   t[3580] := 1_070_001_024;
   t[3581] := 1_070_002_013;
   t[3582] := 1_070_003_096;
   t[3583] := 2_071_201_008;
   t[3584] := 2_071_202_005;
   t[3585] := 2_071_403_104;
   t[3586] := 71403105;
   t[3587] := 71502007;
   t[3588] := 71503043;
   t[3589] := 1_071_501_000;
   t[3590] := 1_071_502_003;
   t[3591] := 73603047;
   t[3592] := 2_073_602_002;
   t[3593] := 73602000;
   t[3594] := 73603013;
   t[3595] := 83001002;
   t[3596] := 1_083_001_014;
   t[3597] := 1_083_002_004;
   t[3598] := 1_084_801_030;
   t[3599] := 1_084_802_012;
   t[3600] := 2_084_801_022;
   t[3601] := 2_084_802_008;
   t[3602] := 84801020;
   t[3603] := 1_084_801_016;
   t[3604] := 85001000;
   t[3605] := 85002000;
   t[3606] := 2_085_101_016;
   t[3607] := 2_085_102_008;
   t[3608] := 1_086_312_107;
   t[3609] := 2_089_703_009;
   t[3610] := 2_090_203_001;
   t[3611] := 90203000;
   t[3612] := 94102009;
   t[3613] := 1_094_101_024;
   t[3614] := 1_094_102_013;
   t[3615] := 1_094_103_096;
   t[3616] := 1_095_201_008;
   t[3617] := 1_095_202_005;
   t[3618] := 2_095_403_104;
   t[3619] := 95403105;
   t[3620] := 95502007;
   t[3621] := 95503043;
   t[3622] := 1_095_501_000;
   t[3623] := 1_095_502_003;
   t[3624] := 97603047;
   t[3625] := 2_097_602_002;
   t[3626] := 97602000;
   t[3627] := 97603013;
   t[3628] := 1_110_312_108;
   t[3629] := 2_113_803_009;
   t[3630] := 114_303_001;
   t[3631] := 1_114_303_000;
   t[3632] := 148_701_002;
   t[3633] := 1_148_701_014;
   t[3634] := 1_148_702_004;
   t[3635] := 150_501_030;
   t[3636] := 150_502_012;
   t[3637] := 1_150_501_022;
   t[3638] := 1_150_502_008;
   t[3639] := 2_150_501_020;
   t[3640] := 150_501_016;
   t[3641] := 150_701_000;
   t[3642] := 150_702_000;
   t[3643] := 150_801_016;
   t[3644] := 150_802_008;
   t[3645] := 1_151_101_000;
   t[3646] := 1_151_102_000;
   t[3647] := 1_151_101_016;
   t[3648] := 1_151_102_008;
   t[3649] := 2_153_502_009;
   t[3650] := 153_501_024;
   t[3651] := 153_502_013;
   t[3652] := 153_503_096;
   t[3653] := 1_154_001_008;
   t[3654] := 1_154_002_005;
   t[3655] := 2_154_101_024;
   t[3656] := 2_154_102_013;
   t[3657] := 2_154_301_008;
   t[3658] := 2_154_302_005;
   t[3659] := 2_154_401_024;
   t[3660] := 2_154_402_013;
   t[3661] := 2_154_601_008;
   t[3662] := 2_154_602_005;
   t[3663] := 154_903_104;
   t[3664] := 1_154_903_105;
   t[3665] := 155_002_007;
   t[3666] := 155_003_043;
   t[3667] := 1_155_001_000;
   t[3668] := 1_155_002_003;
   t[3669] := 2_157_003_047;
   t[3670] := 1_157_002_002;
   t[3671] := 2_157_002_000;
   t[3672] := 2_157_003_013;
   t[3673] := 170_012_109;
   t[3674] := 2_173_703_009;
   t[3675] := 2_174_103_001;
   t[3676] := 174_103_000;
   t[3677] := 269_401_002;
   t[3678] := 1_269_401_014;
   t[3679] := 1_269_402_004;
   t[3680] := 271_101_030;
   t[3681] := 271_102_012;
   t[3682] := 1_271_101_022;
   t[3683] := 1_271_102_008;
   t[3684] := 2_271_101_020;
   t[3685] := 271_101_016;
   t[3686] := 1_271_301_000;
   t[3687] := 1_271_302_000;
   t[3688] := 2_271_401_016;
   t[3689] := 2_271_402_008;
   t[3690] := 274_102_009;
   t[3691] := 1_274_101_024;
   t[3692] := 1_274_102_013;
   t[3693] := 1_274_103_096;
   t[3694] := 2_275_101_008;
   t[3695] := 2_275_102_005;
   t[3696] := 1_275_403_104;
   t[3697] := 2_275_403_105;
   t[3698] := 1_275_402_007;
   t[3699] := 1_275_403_043;
   t[3700] := 2_275_401_000;
   t[3701] := 2_275_402_003;
   t[3702] := 2_277_403_047;
   t[3703] := 1_277_402_002;
   t[3704] := 2_277_402_000;
   t[3705] := 2_277_403_013;
   t[3706] := 1_290_212_110;
   t[3707] := 2_294_103_009;
   t[3708] := 294_303_001;
   t[3709] := 1_294_303_000;
   t[3710] := 380_401_002;
   t[3711] := 1_380_401_014;
   t[3712] := 1_380_402_004;
   t[3713] := 2_382_301_030;
   t[3714] := 2_382_302_012;
   t[3715] := 382_301_022;
   t[3716] := 382_302_008;
   t[3717] := 1_382_301_020;
   t[3718] := 2_382_301_016;
   t[3719] := 382_501_000;
   t[3720] := 382_502_000;
   t[3721] := 2_382_601_016;
   t[3722] := 2_382_602_008;
   t[3723] := 1_385_202_009;
   t[3724] := 2_385_201_024;
   t[3725] := 2_385_202_013;
   t[3726] := 2_385_203_096;
   t[3727] := 2_386_301_008;
   t[3728] := 2_386_302_005;
   t[3729] := 386_503_104;
   t[3730] := 1_386_503_105;
   t[3731] := 386_602_007;
   t[3732] := 386_603_043;
   t[3733] := 1_386_601_000;
   t[3734] := 1_386_602_003;
   t[3735] := 1_388_803_047;
   t[3736] := 388_802_002;
   t[3737] := 1_388_802_000;
   t[3738] := 1_388_803_013;
   t[3739] := 2_401_612_111;
   t[3740] := 405_503_009;
   t[3741] := 405_803_001;
   t[3742] := 1_405_803_000;
   t[3743] := 410_103_008;
   t[3744] := 1_410_103_009;
   t[3745] := 410_403_013;
   t[3746] := 417_003_029;
   t[3747] := 1_417_003_189;
   t[3748] := 2_417_503_185;
   t[3749] := 417_601_002;
   t[3750] := 1_417_601_014;
   t[3751] := 1_417_602_004;
   t[3752] := 1_418_103_189;
   t[3753] := 1_418_303_181;
   t[3754] := 418_303_177;
   t[3755] := 1_418_303_176;
   t[3756] := 2_418_803_180;
   t[3757] := 418_903_181;
   t[3758] := 1_419_003_177;
   t[3759] := 2_419_103_176;
   t[3760] := 2_419_501_030;
   t[3761] := 2_419_502_012;
   t[3762] := 419_501_022;
   t[3763] := 419_502_008;
   t[3764] := 1_419_501_020;
   t[3765] := 2_419_501_016;
   t[3766] := 2_419_801_000;
   t[3767] := 2_419_802_000;
   t[3768] := 419_801_016;
   t[3769] := 419_802_008;
   t[3770] := 1_421_603_160;
   t[3771] := 2_421_603_000;
   t[3772] := 1_425_612_112;
   t[3773] := 1_426_803_008;
   t[3774] := 2_426_803_009;
   t[3775] := 1_427_503_001;
   t[3776] := 2_427_503_000;
   t[3777] := 2_431_002_009;
   t[3778] := 431_001_024;
   t[3779] := 431_002_013;
   t[3780] := 431_003_096;
   t[3781] := 2_432_001_008;
   t[3782] := 2_432_002_005;
   t[3783] := 432_303_104;
   t[3784] := 1_432_303_105;
   t[3785] := 1_432_402_007;
   t[3786] := 1_432_403_043;
   t[3787] := 2_432_401_000;
   t[3788] := 2_432_402_003;
   t[3789] := 2_434_503_047;
   t[3790] := 1_434_502_002;
   t[3791] := 2_434_502_000;
   t[3792] := 2_434_503_013;
   t[3793] := 1_434_501_002;
   t[3794] := 2_434_501_014;
   t[3795] := 2_434_502_004;
   t[3796] := 2_436_401_030;
   t[3797] := 2_436_402_012;
   t[3798] := 436_401_022;
   t[3799] := 436_402_008;
   t[3800] := 1_436_401_020;
   t[3801] := 2_436_401_016;
   t[3802] := 447_212_113;
   t[3803] := 2_450_003_009;
   t[3804] := 2_450_403_001;
   t[3805] := 450_403_000;
   t[3806] := 2_454_302_009;
   t[3807] := 454_301_024;
   t[3808] := 454_302_013;
   t[3809] := 454_303_096;
   t[3810] := 2_455_501_008;
   t[3811] := 2_455_502_005;
   t[3812] := 455_803_104;
   t[3813] := 1_455_803_105;
   t[3814] := 455_802_007;
   t[3815] := 455_803_043;
   t[3816] := 1_455_901_000;
   t[3817] := 1_455_902_003;
   t[3818] := 1_458_003_047;
   t[3819] := 458_002_002;
   t[3820] := 1_458_002_000;
   t[3821] := 1_458_003_013;
   t[3822] := 1_470_712_114;
   t[3823] := 2_473_703_009;
   t[3824] := 474_003_001;
   t[3825] := 1_474_003_000;
   t[3826] := 1_548_401_002;
   t[3827] := 2_548_401_014;
   t[3828] := 2_548_402_004;
   t[3829] := 1_550_301_030;
   t[3830] := 1_550_302_012;
   t[3831] := 2_550_301_022;
   t[3832] := 2_550_302_008;
   t[3833] := 550_301_020;
   t[3834] := 1_550_301_016;
   t[3835] := 2_550_601_000;
   t[3836] := 2_550_602_000;
   t[3837] := 550_601_016;
   t[3838] := 550_602_008;
   t[3839] := 2_553_202_009;
   t[3840] := 553_201_024;
   t[3841] := 553_202_013;
   t[3842] := 553_203_096;
   t[3843] := 1_554_401_008;
   t[3844] := 1_554_402_005;
   t[3845] := 2_554_703_104;
   t[3846] := 554_703_105;
   t[3847] := 2_554_702_007;
   t[3848] := 2_554_703_043;
   t[3849] := 554_701_000;
   t[3850] := 554_702_003;
   t[3851] := 1_556_903_047;
   t[3852] := 557_002_002;
   t[3853] := 1_557_002_000;
   t[3854] := 1_557_003_013;
   t[3855] := 569_712_115;
   t[3856] := 2_572_703_009;
   t[3857] := 1_573_103_001;
   t[3858] := 2_573_103_000;
   t[3859] := 1_616_813_011;
   t[3860] := 1_620_201_002;
   t[3861] := 2_620_201_014;
   t[3862] := 2_620_202_004;
   t[3863] := 2_622_001_030;
   t[3864] := 2_622_002_012;
   t[3865] := 622_001_022;
   t[3866] := 622_002_008;
   t[3867] := 1_622_001_020;
   t[3868] := 2_622_001_016;
   t[3869] := 622_101_000;
   t[3870] := 622_102_000;
   t[3871] := 1_622_201_016;
   t[3872] := 1_622_202_008;
   t[3873] := 624_902_009;
   t[3874] := 1_624_901_024;
   t[3875] := 1_624_902_013;
   t[3876] := 1_624_903_096;
   t[3877] := 1_626_001_008;
   t[3878] := 1_626_002_005;
   t[3879] := 626_303_104;
   t[3880] := 1_626_303_105;
   t[3881] := 626_402_007;
   t[3882] := 626_403_043;
   t[3883] := 1_626_401_000;
   t[3884] := 1_626_402_003;
   t[3885] := 2_628_503_047;
   t[3886] := 628_513_012;
   t[3887] := 1_628_502_002;
   t[3888] := 2_628_502_000;
   t[3889] := 2_628_503_013;
   t[3890] := 1_630_913_013;
   t[3891] := 635_413_014;
   t[3892] := 1_637_413_015;
   t[3893] := 641_313_016;
   t[3894] := 1_641_312_116;
   t[3895] := 2_644_403_009;
   t[3896] := 2_644_603_001;
   t[3897] := 644_703_000;
   t[3898] := 2_647_013_010;
   t[3899] := 647_013_011;
   t[3900] := 1_687_101_002;
   t[3901] := 2_687_101_014;
   t[3902] := 2_687_102_004;
   t[3903] := 688_901_030;
   t[3904] := 688_902_012;
   t[3905] := 1_688_901_022;
   t[3906] := 1_688_902_008;
   t[3907] := 2_688_901_020;
   t[3908] := 688_901_016;
   t[3909] := 689_001_000;
   t[3910] := 689_002_000;
   t[3911] := 2_689_201_016;
   t[3912] := 2_689_202_008;
   t[3913] := 2_691_902_009;
   t[3914] := 691_901_024;
   t[3915] := 691_902_013;
   t[3916] := 691_903_096;
   t[3917] := 693_001_008;
   t[3918] := 693_002_005;
   t[3919] := 693_303_104;
   t[3920] := 1_693_303_105;
   t[3921] := 1_693_402_007;
   t[3922] := 1_693_403_043;
   t[3923] := 2_693_401_000;
   t[3924] := 2_693_402_003;
   t[3925] := 1_695_503_047;
   t[3926] := 2_695_513_012;
   t[3927] := 695_502_002;
   t[3928] := 1_695_502_000;
   t[3929] := 1_695_503_013;
   t[3930] := 1_697_913_013;
   t[3931] := 702_413_014;
   t[3932] := 704_413_015;
   t[3933] := 708_313_016;
   t[3934] := 1_708_312_117;
   t[3935] := 2_711_403_009;
   t[3936] := 1_711_703_001;
   t[3937] := 2_711_703_000;
   t[3938] := 2_714_013_010;
   t[3939] := 714_013_011;
   t[3940] := 1_980_801_002;
   t[3941] := 2_980_801_014;
   t[3942] := 2_980_802_004;
   t[3943] := 1_982_601_030;
   t[3944] := 1_982_602_012;
   t[3945] := 2_982_601_022;
   t[3946] := 2_982_602_008;
   t[3947] := 982_601_020;
   t[3948] := 1_982_601_016;
   t[3949] := 982_701_000;
   t[3950] := 982_702_000;
   t[3951] := 982_901_016;
   t[3952] := 982_902_008;
   t[3953] := 2_985_602_009;
   t[3954] := 985_601_024;
   t[3955] := 985_602_013;
   t[3956] := 985_603_096;
   t[3957] := 986_601_008;
   t[3958] := 986_602_005;
   t[3959] := 2_986_903_104;
   t[3960] := 986_903_105;
   t[3961] := 987_002_007;
   t[3962] := 987_003_043;
   t[3963] := 1_987_001_000;
   t[3964] := 1_987_002_003;
   t[3965] := 2_988_903_047;
   t[3966] := 988_913_012;
   t[3967] := 1_988_902_002;
   t[3968] := 2_988_902_000;
   t[3969] := 2_988_903_013;
   t[3970] := 991_213_013;
   t[3971] := 1_995_613_014;
   t[3972] := 1_997_513_015;
   t[3973] := 60911;
   t[3974] := 501002;
   t[3975] := 1_000_601_014;
   t[3976] := 1_000_602_004;
   t[3977] := 1413016;
   t[3978] := 1_001_412_118;
   t[3979] := 2_002_201_030;
   t[3980] := 2_002_202_012;
   t[3981] := 2301022;
   t[3982] := 2302008;
   t[3983] := 1_002_301_020;
   t[3984] := 2_002_301_016;
   t[3985] := 1_004_603_009;
   t[3986] := 2_004_903_001;
   t[3987] := 4903000;
   t[3988] := 1_007_113_010;
   t[3989] := 2_007_113_011;
   t[3990] := 2_008_802_009;
   t[3991] := 8801024;
   t[3992] := 8802013;
   t[3993] := 8803096;
   t[3994] := 2_009_801_008;
   t[3995] := 2_009_802_005;
   t[3996] := 2_010_103_104;
   t[3997] := 10103105;
   t[3998] := 1_010_102_007;
   t[3999] := 1_010_103_043;
   t[4000] := 2_010_201_000;
   t[4001] := 2_010_202_003;
   t[4002] := 12103047;
   t[4003] := 1_012_113_012;
   t[4004] := 2_012_102_002;
   t[4005] := 12102000;
   t[4006] := 12103013;
   t[4007] := 2_014_413_013;
   t[4008] := 2_018_913_014;
   t[4009] := 1_020_813_015;
   t[4010] := 2_024_713_016;
   t[4011] := 24712119;
   t[4012] := 1_027_803_009;
   t[4013] := 1_028_203_001;
   t[4014] := 2_028_203_000;
   t[4015] := 2_030_413_010;
   t[4016] := 30413011;
   t[4017] := 1_048_201_002;
   t[4018] := 2_048_201_014;
   t[4019] := 2_048_202_004;
   t[4020] := 1_050_101_030;
   t[4021] := 1_050_102_012;
   t[4022] := 2_050_101_022;
   t[4023] := 2_050_102_008;
   t[4024] := 50101020;
   t[4025] := 1_050_101_016;
   t[4026] := 2_050_201_000;
   t[4027] := 2_050_202_000;
   t[4028] := 1_050_401_016;
   t[4029] := 1_050_402_008;
   t[4030] := 1_053_002_009;
   t[4031] := 2_053_001_024;
   t[4032] := 2_053_002_013;
   t[4033] := 2_053_003_096;
   t[4034] := 54101008;
   t[4035] := 54102005;
   t[4036] := 1_054_303_104;
   t[4037] := 2_054_303_105;
   t[4038] := 2_054_402_007;
   t[4039] := 2_054_403_043;
   t[4040] := 54401000;
   t[4041] := 54402003;
   t[4042] := 2_056_303_047;
   t[4043] := 56313012;
   t[4044] := 1_056_302_002;
   t[4045] := 2_056_302_000;
   t[4046] := 2_056_303_013;
   t[4047] := 2_058_613_013;
   t[4048] := 2_063_013_014;
   t[4049] := 1_065_013_015;
   t[4050] := 1_068_913_016;
   t[4051] := 2_068_912_120;
   t[4052] := 69901002;
   t[4053] := 1_069_901_014;
   t[4054] := 1_069_902_004;
   t[4055] := 71801030;
   t[4056] := 71802012;
   t[4057] := 1_071_801_022;
   t[4058] := 1_071_802_008;
   t[4059] := 2_071_801_020;
   t[4060] := 71801016;
   t[4061] := 1_072_103_009;
   t[4062] := 72403001;
   t[4063] := 1_072_403_000;
   t[4064] := 2_074_613_010;
   t[4065] := 74613011;
   t[4066] := 1_076_302_009;
   t[4067] := 2_076_301_024;
   t[4068] := 2_076_302_013;
   t[4069] := 2_076_303_096;
   t[4070] := 2_077_401_008;
   t[4071] := 2_077_402_005;
   t[4072] := 2_077_703_104;
   t[4073] := 77703105;
   t[4074] := 77802007;
   t[4075] := 77803043;
   t[4076] := 1_077_801_000;
   t[4077] := 1_077_802_003;
   t[4078] := 2_079_903_047;
   t[4079] := 79913012;
   t[4080] := 1_079_902_002;
   t[4081] := 2_080_002_000;
   t[4082] := 2_080_003_013;
   t[4083] := 82213013;
   t[4084] := 86813014;
   t[4085] := 1_088_713_015;
   t[4086] := 1_097_313_001;
   t[4087] := 1_464_303_005;
   t[4088] := 1_464_603_013;
   t[4089] := 483_113_000;
   t[4090] := 2_484_313_010;
   t[4091] := 1_484_313_001;
   t[4092] := 519_503_005;
   t[4093] := 1_519_803_013;
   t[4094] := 520_003_009;
   t[4095] := 1_521_603_001;
   t[4096] := 2_521_603_000;
   t[4097] := 526_613_000;
   t[4098] := 1_527_113_010;
   t[4099] := 2_527_113_011;
   t[4100] := 535_801_002;
   t[4101] := 1_535_801_014;
   t[4102] := 1_535_802_004;
   t[4103] := 2_537_701_030;
   t[4104] := 2_537_702_012;
   t[4105] := 537_701_022;
   t[4106] := 537_702_008;
   t[4107] := 1_537_701_020;
   t[4108] := 2_537_701_016;
   t[4109] := 1_537_901_000;
   t[4110] := 1_537_902_000;
   t[4111] := 2_538_001_016;
   t[4112] := 2_538_002_008;
   t[4113] := 2_540_803_004;
   t[4114] := 540_803_005;
   t[4115] := 540_903_001;
   t[4116] := 1_540_903_000;
   t[4117] := 2_541_703_008;
   t[4118] := 541_703_009;
   t[4119] := 2_541_803_001;
   t[4120] := 541_803_000;
   t[4121] := 2_557_402_024;
   t[4122] := 2_557_402_025;
   t[4123] := 557_401_024;
   t[4124] := 557_402_029;
   t[4125] := 557_403_096;
   t[4126] := 558_501_008;
   t[4127] := 558_502_021;
   t[4128] := 2_558_703_104;
   t[4129] := 558_703_105;
   t[4130] := 1_558_802_023;
   t[4131] := 1_558_803_043;
   t[4132] := 2_558_801_000;
   t[4133] := 2_558_802_019;
   t[4134] := 1_558_902_018;
   t[4135] := 2_558_902_016;
   t[4136] := 2_558_903_009;
   t[4137] := 1_580_503_013;
   t[4138] := 1_580_513_012;
   t[4139] := 2_582_813_013;
   t[4140] := 2_587_313_014;
   t[4141] := 1_589_213_015;
   t[4142] := 1_593_013_016;
   t[4143] := 2_593_012_121;
   t[4144] := 596_503_009;
   t[4145] := 1_596_803_001;
   t[4146] := 2_596_803_000;
   t[4147] := 2_598_913_010;
   t[4148] := 598_913_011;
   t[4149] := 1_634_201_002;
   t[4150] := 2_634_201_014;
   t[4151] := 2_634_202_020;
   t[4152] := 636_101_030;
   t[4153] := 636_102_028;
   t[4154] := 1_636_101_022;
   t[4155] := 1_636_102_024;
   t[4156] := 2_636_101_020;
   t[4157] := 636_101_016;
   t[4158] := 1_636_301_000;
   t[4159] := 1_636_302_016;
   t[4160] := 636_301_016;
   t[4161] := 636_302_024;
   t[4162] := 636_401_000;
   t[4163] := 636_402_016;
   t[4164] := 636_401_016;
   t[4165] := 636_402_024;
   t[4166] := 2_639_102_025;
   t[4167] := 639_101_024;
   t[4168] := 639_102_029;
   t[4169] := 639_103_096;
   t[4170] := 1_640_201_008;
   t[4171] := 1_640_202_021;
   t[4172] := 640_503_104;
   t[4173] := 1_640_503_105;
   t[4174] := 640_502_023;
   t[4175] := 640_503_043;
   t[4176] := 1_640_501_000;
   t[4177] := 1_640_502_019;
   t[4178] := 1_642_502_003;
   t[4179] := 1_642_503_047;
   t[4180] := 2_642_513_012;
   t[4181] := 642_502_002;
   t[4182] := 1_642_602_000;
   t[4183] := 1_642_603_013;
   t[4184] := 1_644_813_013;
   t[4185] := 649_213_014;
   t[4186] := 651_213_015;
   t[4187] := 655_113_016;
   t[4188] := 1_655_112_122;
   t[4189] := 1_658_403_009;
   t[4190] := 1_658_803_001;
   t[4191] := 2_658_803_000;
   t[4192] := 2_661_013_010;
   t[4193] := 661_013_011;
   t[4194] := 2_662_702_016;
   t[4195] := 2_975_801_002;
   t[4196] := 975_801_014;
   t[4197] := 975_802_020;
   t[4198] := 977_501_030;
   t[4199] := 977_502_028;
   t[4200] := 1_977_501_022;
   t[4201] := 1_977_502_024;
   t[4202] := 2_977_601_020;
   t[4203] := 977_601_016;
   t[4204] := 977_701_000;
   t[4205] := 977_702_016;
   t[4206] := 2_977_801_016;
   t[4207] := 2_977_802_024;
   t[4208] := 2_980_402_025;
   t[4209] := 980_401_024;
   t[4210] := 980_402_029;
   t[4211] := 980_403_096;
   t[4212] := 1_981_201_008;
   t[4213] := 1_981_202_021;
   t[4214] := 1_981_301_024;
   t[4215] := 1_981_302_029;
   t[4216] := 981_301_008;
   t[4217] := 981_302_021;
   t[4218] := 2_981_301_024;
   t[4219] := 2_981_302_029;
   t[4220] := 981_501_008;
   t[4221] := 981_502_021;
   t[4222] := 981_703_104;
   t[4223] := 1_981_703_105;
   t[4224] := 2_981_802_023;
   t[4225] := 2_981_803_043;
   t[4226] := 981_801_000;
   t[4227] := 981_802_019;
   t[4228] := 2_982_003_035;
   t[4229] := 982_103_043;
   t[4230] := 2_983_802_003;
   t[4231] := 2_983_803_047;
   t[4232] := 983_813_012;
   t[4233] := 1_983_802_002;
   t[4234] := 2_983_802_000;
   t[4235] := 2_983_803_013;
   t[4236] := 1_986_013_013;
   t[4237] := 1_990_713_014;
   t[4238] := 992_613_015;
   t[4239] := 1_996_513_016;
   t[4240] := 2_996_512_123;
   t[4241] := 60930;
   t[4242] := 2_000_103_009;
   t[4243] := 2_000_403_001;
   t[4244] := 403000;
   t[4245] := 2513010;
   t[4246] := 1_002_513_011;
   t[4247] := 2_004_102_016;
   t[4248] := 44301002;
   t[4249] := 1_044_301_014;
   t[4250] := 1_044_302_020;
   t[4251] := 46101030;
   t[4252] := 46102028;
   t[4253] := 1_046_101_022;
   t[4254] := 1_046_102_024;
   t[4255] := 2_046_101_020;
   t[4256] := 46101016;
   t[4257] := 1_046_201_000;
   t[4258] := 1_046_202_016;
   t[4259] := 1_046_401_016;
   t[4260] := 1_046_402_024;
   t[4261] := 1_049_102_025;
   t[4262] := 2_049_101_024;
   t[4263] := 2_049_102_029;
   t[4264] := 2_049_103_096;
   t[4265] := 50101008;
   t[4266] := 50102021;
   t[4267] := 2_050_403_104;
   t[4268] := 50403105;
   t[4269] := 1_050_502_023;
   t[4270] := 1_050_503_043;
   t[4271] := 2_050_501_000;
   t[4272] := 2_050_502_019;
   t[4273] := 1_052_502_003;
   t[4274] := 1_052_503_047;
   t[4275] := 2_052_513_012;
   t[4276] := 52502002;
   t[4277] := 1_052_502_000;
   t[4278] := 1_052_503_013;
   t[4279] := 54813013;
   t[4280] := 1_059_213_014;
   t[4281] := 1_061_213_015;
   t[4282] := 2_065_013_016;
   t[4283] := 65012124;
   t[4284] := 1_068_603_009;
   t[4285] := 2_068_903_001;
   t[4286] := 68903000;
   t[4287] := 2_071_113_010;
   t[4288] := 71213011;
   t[4289] := 1_072_802_016;
   t[4290] := 123_213_017;
   t[4291] := 124_902_000;
   t[4292] := 124_903_008;
   t[4293] := 1_124_903_009;
   t[4294] := 1_125_103_013;
   t[4295] := 127_213_018;
   t[4296] := 1_131_603_029;
   t[4297] := 2_131_603_189;
   t[4298] := 2_131_610_001;
   t[4299] := 2_131_611_124;
   t[4300] := 2_131_613_000;
   t[4301] := 132_003_185;
   t[4302] := 132_703_189;
   t[4303] := 132_803_185;
   t[4304] := 1_132_803_177;
   t[4305] := 2_132_903_176;
   t[4306] := 133_503_180;
   t[4307] := 1_133_503_181;
   t[4308] := 133_603_177;
   t[4309] := 1_133_603_176;
   t[4310] := 136_103_160;
   t[4311] := 1_136_103_000;
   t[4312] := 1_136_113_010;
   t[4313] := 2_136_113_015;
   t[4314] := 2_140_013_016;
   t[4315] := 140_012_125;
   t[4316] := 2_141_303_008;
   t[4317] := 141_303_009;
   t[4318] := 141_903_001;
   t[4319] := 1_141_903_000;
   t[4320] := 1_145_313_010;
   t[4321] := 2_145_313_011;
   t[4322] := 145_302_016;
   t[4323] := 1_150_713_000;
   t[4324] := 0;
   t[4325] := 0;
   t[4326] := 0;
   t[4327] := 0;
   t[4328] := 0;
   t[4329] := 0;
   t[4330] := 0;
   t[4331] := 0;
   t[4332] := 0;
   t[4333] := 0;
   t[4334] := 0;
   t[4335] := 0;
   t[4336] := 0;
   t[4337] := 0;
   t[4338] := 0;
   t[4339] := 0;
   t[4340] := 0;
   t[4341] := 0;
   t[4342] := 0;
   t[4343] := 0;
   t[4344] := 0;
   t[4345] := 0;
   t[4346] := 0;
   t[4347] := 0;
   t[4348] := 0;
   t[4349] := 0;
   t[4350] := 0;
   t[4351] := 0;
   t[4352] := 0;
   t[4353] := 0;
   t[4354] := 0;
   t[4355] := 0;
   t[4356] := 0;
   t[4357] := 0;
   t[4358] := 0;
   t[4359] := 0;
   t[4360] := 0;
   t[4361] := 0;
   t[4362] := 0;
   t[4363] := 0;
   t[4364] := 0;
   t[4365] := 0;
   t[4366] := 0;
   t[4367] := 0;
   t[4368] := 0;
   t[4369] := 0;
   t[4370] := 0;
   t[4371] := 0;
   t[4372] := 0;
   t[4373] := 0;
   t[4374] := 0;
   t[4375] := 0;
   t[4376] := 0;
   t[4377] := 0;
   t[4378] := 0;
   t[4379] := 0;
   t[4380] := 0;
   t[4381] := 0;
   t[4382] := 0;
   t[4383] := 0;
   t[4384] := 0;
   t[4385] := 0;
   t[4386] := 0;
   t[4387] := 0;
   t[4388] := 0;
   t[4389] := 0;
   t[4390] := 0;
   t[4391] := 0;
   t[4392] := 0;
   t[4393] := 0;
   t[4394] := 0;
   t[4395] := 0;
   t[4396] := 0;
   t[4397] := 0;
   t[4398] := 0;
   t[4399] := 0;
   t[4400] := 0;
   t[4401] := 0;
   t[4402] := 0;
   t[4403] := 0;
   t[4404] := 0;
   t[4405] := 0;
   t[4406] := 0;
   t[4407] := 0;
   t[4408] := 0;
   t[4409] := 0;
   t[4410] := 0;
   t[4411] := 0;
   t[4412] := 0;
   t[4413] := 0;
   t[4414] := 0;
   t[4415] := 0;
   t[4416] := 0;
   t[4417] := 0;
   t[4418] := 0;
   t[4419] := 0;
   t[4420] := 0;
   t[4421] := 0;
   t[4422] := 0;
   t[4423] := 0;
   t[4424] := 0;
   t[4425] := 0;
   t[4426] := 0;
   t[4427] := 0;
   t[4428] := 0;
   t[4429] := 0;
   t[4430] := 0;
   t[4431] := 0;
   t[4432] := 0;
   t[4433] := 0;
   t[4434] := 0;
   t[4435] := 0;
   t[4436] := 0;
   t[4437] := 0;
   t[4438] := 0;
   t[4439] := 0;
   t[4440] := 0;
   t[4441] := 0;
   t[4442] := 0;
   t[4443] := 0;
   t[4444] := 0;
   t[4445] := 0;
   t[4446] := 0;
   t[4447] := 0;
   t[4448] := 0;
   t[4449] := 0;
   t[4450] := 0;
   t[4451] := 0;
   t[4452] := 0;
   t[4453] := 0;
   t[4454] := 0;
   t[4455] := 0;
   t[4456] := 0;
   t[4457] := 0;
   t[4458] := 0;
   t[4459] := 0;
   t[4460] := 0;
   t[4461] := 0;
   t[4462] := 0;
   t[4463] := 0;
   t[4464] := 0;
   t[4465] := 0;
   t[4466] := 0;
   t[4467] := 0;
   t[4468] := 0;
   t[4469] := 0;
   t[4470] := 0;
   t[4471] := 0;
   t[4472] := 0;
   t[4473] := 0;
   t[4474] := 0;
   t[4475] := 0;
   t[4476] := 0;
   t[4477] := 0;
   t[4478] := 0;
   t[4479] := 0;
   t[4480] := 0;
   t[4481] := 0;
   t[4482] := 0;
   t[4483] := 0;
   t[4484] := 0;
   t[4485] := 0;
   t[4486] := 0;
   t[4487] := 0;
   t[4488] := 0;
   t[4489] := 0;
   t[4490] := 0;
   t[4491] := 0;
   t[4492] := 0;
   t[4493] := 0;
   t[4494] := 0;
   t[4495] := 0;
   t[4496] := 0;
   t[4497] := 0;
   t[4498] := 0;
   t[4499] := 0;
   t[4500] := 0;
   t[4501] := 0;
   t[4502] := 0;
   t[4503] := 0;
   t[4504] := 0;
   t[4505] := 0;
   t[4506] := 0;
   t[4507] := 0;
   t[4508] := 0;
   t[4509] := 0;
   t[4510] := 0;
   t[4511] := 0;
   t[4512] := 0;
   t[4513] := 0;
   t[4514] := 0;
   t[4515] := 0;
   t[4516] := 0;
   t[4517] := 0;
   t[4518] := 0;
   t[4519] := 0;
   t[4520] := 0;
   t[4521] := 0;
   t[4522] := 0;
   t[4523] := 0;
   t[4524] := 0;
   t[4525] := 0;
   t[4526] := 0;
   t[4527] := 0;
   t[4528] := 0;
   t[4529] := 0;
   t[4530] := 0;
   t[4531] := 0;
   t[4532] := 0;
   t[4533] := 0;
   t[4534] := 0;
   t[4535] := 0;
   t[4536] := 0;
   t[4537] := 0;
   t[4538] := 0;
   t[4539] := 0;
   t[4540] := 0;
   t[4541] := 0;
   t[4542] := 0;
   t[4543] := 0;
   t[4544] := 0;
   t[4545] := 0;
   t[4546] := 0;
   t[4547] := 0;
   t[4548] := 0;
   t[4549] := 0;
   t[4550] := 0;
   t[4551] := 0;
   t[4552] := 0;
   t[4553] := 0;
   t[4554] := 0;
   t[4555] := 0;
   t[4556] := 0;
   t[4557] := 0;
   t[4558] := 0;
   t[4559] := 0;
   t[4560] := 0;
   t[4561] := 0;
   t[4562] := 0;
   t[4563] := 0;
   t[4564] := 0;
   t[4565] := 0;
   t[4566] := 0;
   t[4567] := 0;
   t[4568] := 0;
   t[4569] := 0;
   t[4570] := 0;
   t[4571] := 0;
   t[4572] := 0;
   t[4573] := 0;
   t[4574] := 0;
   t[4575] := 0;
   t[4576] := 0;
   t[4577] := 0;
   t[4578] := 0;
   t[4579] := 0;
   t[4580] := 0;
   t[4581] := 0;
   t[4582] := 0;
   t[4583] := 0;
   t[4584] := 0;
   t[4585] := 0;
   t[4586] := 0;
   t[4587] := 0;
   t[4588] := 0;
   t[4589] := 0;
   t[4590] := 0;
   t[4591] := 0;
   t[4592] := 0;
   t[4593] := 0;
   t[4594] := 0;
   t[4595] := 0;
   t[4596] := 0;
   t[4597] := 0;
   t[4598] := 0;
   t[4599] := 0;
   t[4600] := 0;
   t[4601] := 0;
   t[4602] := 0;
   t[4603] := 0;
   t[4604] := 0;
   t[4605] := 0;
   t[4606] := 0;
   t[4607] := 0;
   t[4608] := 0;
   t[4609] := 0;
   t[4610] := 0;
   t[4611] := 0;
   t[4612] := 0;
   t[4613] := 0;
   t[4614] := 0;
   t[4615] := 0;
   t[4616] := 0;
   t[4617] := 0;
   t[4618] := 0;
   t[4619] := 0;
   t[4620] := 0;
   t[4621] := 0;
   t[4622] := 0;
   t[4623] := 0;
   t[4624] := 0;
   t[4625] := 0;
   t[4626] := 0;
   t[4627] := 0;
   t[4628] := 0;
   t[4629] := 0;
   t[4630] := 0;
   t[4631] := 0;
   t[4632] := 0;
   t[4633] := 0;
   t[4634] := 0;
   t[4635] := 0;
   t[4636] := 0;
   t[4637] := 0;
   t[4638] := 0;
   t[4639] := 0;
   t[4640] := 0;
   t[4641] := 0;
   t[4642] := 0;
   t[4643] := 0;
   t[4644] := 0;
   t[4645] := 0;
   t[4646] := 0;
   t[4647] := 0;
   t[4648] := 0;
   t[4649] := 0;
   t[4650] := 0;
   t[4651] := 0;
   t[4652] := 0;
   t[4653] := 0;
   t[4654] := 0;
   t[4655] := 0;
   t[4656] := 0;
   t[4657] := 0;
   t[4658] := 0;
   t[4659] := 0;
   t[4660] := 0;
   t[4661] := 0;
   t[4662] := 0;
   t[4663] := 0;
   t[4664] := 0;
   t[4665] := 0;
   t[4666] := 0;
   t[4667] := 0;
   t[4668] := 0;
   t[4669] := 0;
   t[4670] := 0;
   t[4671] := 0;
   t[4672] := 0;
   t[4673] := 0;
   t[4674] := 0;
   t[4675] := 0;
   t[4676] := 0;
   t[4677] := 0;
   t[4678] := 0;
   t[4679] := 0;
   t[4680] := 0;
   t[4681] := 0;
   t[4682] := 0;
   t[4683] := 0;
   t[4684] := 0;
   t[4685] := 0;
   t[4686] := 0;
   t[4687] := 0;
   t[4688] := 0;
   t[4689] := 0;
   t[4690] := 0;
   t[4691] := 0;
   t[4692] := 0;
   t[4693] := 0;
   t[4694] := 0;
   t[4695] := 0;
   t[4696] := 0;
   t[4697] := 0;
   t[4698] := 0;
   t[4699] := 0;
   t[4700] := 0;
   t[4701] := 0;
   t[4702] := 0;
   t[4703] := 0;
   t[4704] := 0;
   t[4705] := 0;
   t[4706] := 0;
   t[4707] := 0;
   t[4708] := 0;
   t[4709] := 0;
   t[4710] := 0;
   t[4711] := 0;
   t[4712] := 0;
   t[4713] := 0;
   t[4714] := 0;
   t[4715] := 0;
   t[4716] := 0;
   t[4717] := 0;
   t[4718] := 0;
   t[4719] := 0;
   t[4720] := 0;
   t[4721] := 0;
   t[4722] := 0;
   t[4723] := 0;
   t[4724] := 0;
   t[4725] := 0;
   t[4726] := 0;
   t[4727] := 0;
   t[4728] := 0;
   t[4729] := 0;
   t[4730] := 0;
   t[4731] := 0;
   t[4732] := 0;
   t[4733] := 0;
   t[4734] := 0;
   t[4735] := 0;
   t[4736] := 0;
   t[4737] := 0;
   t[4738] := 0;
   t[4739] := 0;
   t[4740] := 0;
   t[4741] := 0;
   t[4742] := 0;
   t[4743] := 0;
   t[4744] := 0;
   t[4745] := 0;
   t[4746] := 0;
   t[4747] := 0;
   t[4748] := 0;
   t[4749] := 0;
   t[4750] := 0;
   t[4751] := 0;
   t[4752] := 0;
   t[4753] := 0;
   t[4754] := 0;
   t[4755] := 0;
   t[4756] := 0;
   t[4757] := 0;
   t[4758] := 0;
   t[4759] := 0;
   t[4760] := 0;
   t[4761] := 0;
   t[4762] := 0;
   t[4763] := 0;
   t[4764] := 0;
   t[4765] := 0;
   t[4766] := 0;
   t[4767] := 0;
   t[4768] := 0;
   t[4769] := 0;
   t[4770] := 0;
   t[4771] := 0;
   t[4772] := 0;
   t[4773] := 0;
   t[4774] := 0;
   t[4775] := 0;
   t[4776] := 0;
   t[4777] := 0;
   t[4778] := 0;
   t[4779] := 0;
   t[4780] := 0;
   t[4781] := 0;
   t[4782] := 0;
   t[4783] := 0;
   t[4784] := 0;
   t[4785] := 0;
   t[4786] := 0;
   t[4787] := 0;
   t[4788] := 0;
   t[4789] := 0;
   t[4790] := 0;
   t[4791] := 0;
   t[4792] := 0;
   t[4793] := 0;
   t[4794] := 0;
   t[4795] := 0;
   t[4796] := 0;
   t[4797] := 0;
   t[4798] := 0;
   t[4799] := 0;
   t[4800] := 0;
   t[4801] := 0;
   t[4802] := 0;
   t[4803] := 0;
   t[4804] := 0;
   t[4805] := 0;
   t[4806] := 0;
   t[4807] := 0;
   t[4808] := 0;
   t[4809] := 0;
   t[4810] := 0;
   t[4811] := 0;
   t[4812] := 0;
   t[4813] := 0;
   t[4814] := 0;
   t[4815] := 0;
   t[4816] := 0;
   t[4817] := 0;
   t[4818] := 0;
   t[4819] := 0;
   t[4820] := 0;
   t[4821] := 0;
   t[4822] := 0;
   t[4823] := 0;
   t[4824] := 0;
   t[4825] := 0;
   t[4826] := 0;
   t[4827] := 0;
   t[4828] := 0;
   t[4829] := 0;
   t[4830] := 0;
   t[4831] := 0;
   t[4832] := 0;
   t[4833] := 0;
   t[4834] := 0;
   t[4835] := 0;
   t[4836] := 0;
   t[4837] := 0;
   t[4838] := 0;
   t[4839] := 0;
   t[4840] := 0;
   t[4841] := 0;
   t[4842] := 0;
   t[4843] := 0;
   t[4844] := 0;
   t[4845] := 0;
   t[4846] := 0;
   t[4847] := 0;
   t[4848] := 0;
   t[4849] := 0;
   t[4850] := 0;
   t[4851] := 0;
   t[4852] := 0;
   t[4853] := 0;
   t[4854] := 0;
   t[4855] := 0;
   t[4856] := 0;
   t[4857] := 0;
   t[4858] := 0;
   t[4859] := 0;
   t[4860] := 0;
   t[4861] := 0;
   t[4862] := 0;
   t[4863] := 0;
   t[4864] := 0;
   t[4865] := 0;
   t[4866] := 0;
   t[4867] := 0;
   t[4868] := 0;
   t[4869] := 0;
   t[4870] := 0;
   t[4871] := 0;
   t[4872] := 0;
   t[4873] := 0;
   t[4874] := 0;
   t[4875] := 0;
   t[4876] := 0;
   t[4877] := 0;
   t[4878] := 0;
   t[4879] := 0;
   t[4880] := 0;
   t[4881] := 0;
   t[4882] := 0;
   t[4883] := 0;
   t[4884] := 0;
   t[4885] := 0;
   t[4886] := 0;
   t[4887] := 0;
   t[4888] := 0;
   t[4889] := 0;
   t[4890] := 0;
   t[4891] := 0;
   t[4892] := 0;
   t[4893] := 0;
   t[4894] := 0;
   t[4895] := 0;
   t[4896] := 0;
   t[4897] := 0;
   t[4898] := 0;
   t[4899] := 0;
   t[4900] := 0;
   t[4901] := 0;
   t[4902] := 0;
   t[4903] := 0;
   t[4904] := 0;
   t[4905] := 0;
   t[4906] := 0;
   t[4907] := 0;
   t[4908] := 0;
   t[4909] := 0;
   t[4910] := 0;
   t[4911] := 0;
   t[4912] := 0;
   t[4913] := 0;
   t[4914] := 0;
   t[4915] := 0;
   t[4916] := 0;
   t[4917] := 0;
   t[4918] := 0;
   t[4919] := 0;
   t[4920] := 0;
   t[4921] := 0;
   t[4922] := 0;
   t[4923] := 0;
   t[4924] := 0;
   t[4925] := 0;
   t[4926] := 0;
   t[4927] := 0;
   t[4928] := 0;
   t[4929] := 0;
   t[4930] := 0;
   t[4931] := 0;
   t[4932] := 0;
   t[4933] := 0;
   t[4934] := 0;
   t[4935] := 0;
   t[4936] := 0;
   t[4937] := 0;
   t[4938] := 0;
   t[4939] := 0;
   t[4940] := 0;
   t[4941] := 0;
   t[4942] := 0;
   t[4943] := 0;
   t[4944] := 0;
   t[4945] := 0;
   t[4946] := 0;
   t[4947] := 0;
   t[4948] := 0;
   t[4949] := 0;
   t[4950] := 0;
   t[4951] := 0;
   t[4952] := 0;
   t[4953] := 0;
   t[4954] := 0;
   t[4955] := 0;
   t[4956] := 0;
   t[4957] := 0;
   t[4958] := 0;
   t[4959] := 0;
   t[4960] := 0;
   t[4961] := 0;
   t[4962] := 0;
   t[4963] := 0;
   t[4964] := 0;
   t[4965] := 0;
   t[4966] := 0;
   t[4967] := 0;
   t[4968] := 0;
   t[4969] := 0;
   t[4970] := 0;
   t[4971] := 0;
   t[4972] := 0;
   t[4973] := 0;
   t[4974] := 0;
   t[4975] := 0;
   t[4976] := 0;
   t[4977] := 0;
   t[4978] := 0;
   t[4979] := 0;
   t[4980] := 0;
   t[4981] := 0;
   t[4982] := 0;
   t[4983] := 0;
   t[4984] := 0;
   t[4985] := 0;
   t[4986] := 0;
   t[4987] := 0;
   t[4988] := 0;
   t[4989] := 0;
   t[4990] := 0;
   t[4991] := 0;
   t[4992] := 0;
   t[4993] := 0;
   t[4994] := 0;
   t[4995] := 0;
   t[4996] := 0;
   t[4997] := 0;
   t[4998] := 0;
   t[4999] := 0;
   t[5000] := 0;
   t[5001] := 0;
   t[5002] := 0;
   t[5003] := 0;
   t[5004] := 0;
   t[5005] := 0;
   t[5006] := 0;
   t[5007] := 0;
   t[5008] := 0;
   t[5009] := 0;
   t[5010] := 0;
   t[5011] := 0;
   t[5012] := 0;
   t[5013] := 0;
   t[5014] := 0;
   t[5015] := 0;
   t[5016] := 0;
   t[5017] := 0;
   t[5018] := 0;
   t[5019] := 0;
   t[5020] := 0;
   t[5021] := 0;
   t[5022] := 0;
   t[5023] := 0;
   t[5024] := 0;
   t[5025] := 0;
   t[5026] := 0;
   t[5027] := 0;
   t[5028] := 0;
   t[5029] := 0;
   t[5030] := 0;
   t[5031] := 0;
   t[5032] := 0;
   t[5033] := 0;
   t[5034] := 0;
   t[5035] := 0;
   t[5036] := 0;
   t[5037] := 0;
   t[5038] := 0;
   t[5039] := 0;
   t[5040] := 0;
   t[5041] := 0;
   t[5042] := 0;
   t[5043] := 0;
   t[5044] := 0;
   t[5045] := 0;
   t[5046] := 0;
   t[5047] := 0;
   t[5048] := 0;
   t[5049] := 0;
   t[5050] := 0;
   t[5051] := 0;
   t[5052] := 0;
   t[5053] := 0;
   t[5054] := 0;
   t[5055] := 0;
   t[5056] := 0;
   t[5057] := 0;